(* Logix 5000 project; controller FV vendor 1 type 14 code 217 rev 31.11; software revision 31.00; part 57 of 63 *)
(* tags used below, declared in another part *)
   CWD : CHECKWORD_FLAGS;
   FV_AV1 : PlantItem;   // AV1
   FV_B42 : INT[255];   // YSVCIP_FLG
   FV_B42_0_2_OutputBit : BOOL;
   FV_B52 : INT[255];   // WASTE_FLG
   FV_N141 : INT[255];   // YSV1 DATA
   FV_N142 : INT[255];   // YSV2 DATA
   FV_N143 : INT[255];   // YSV3 DATA
   FV_N40 : INT[255];   // YSVCIP<PC
   FV_N41 : INT[255];   // YSVCIP>PC
   FV_N50 : INT[255];   // WASTE<PC
   FV_N51 : INT[255];   // WASTE>PC
   FV_T43 : TIMER[10];
   FV_T53 : TIMER[10];
   FV_YSV1R : PlantItem;   // YSV1R
   FV_YSV2O : PlantItem;   // YSV2O
   FV_YSV3O : PlantItem;   // YSV3O
(* FV_Common, continued *)

ROUTINE FV_YSVCIP_CP_21   (* ladder *)
   // Reset command interpreter step counter
   0: XIC(S:FS)CLR(FV_N41[16]);
   // RESET
   1: EQU(FV_N41[16],0)MCR();
   2: OTU(FV_B42[0].0);
   3: OTU(FV_B42[0].1);
   4: OTU(FV_B42[0].8);
   5: FLL(0,FV_N41[0],16);
   // Set PCparameter buffer to 'Null' value
   6: FLL(-32768,FV_N40[1],7);
   7: CLR(FV_N40[0]);
   8: MOV(1,FV_N41[16]);
   9: MCR();
   // ALLOW STARTUP DIALOG
   10: EQU(FV_N41[16],1)MCR();
   // Set process status = ready
   11: MOV(1,FV_N41[0]);
   // Allow startup if any vessel is inactive or on storage control only
   12: [[EQU(FV_N141[0],0) ,EQU(FV_N141[0],5) ] ,[EQU(FV_N142[0],0) ,EQU(FV_N142[0],5) ] ,[EQU(FV_N143[0],0) ,EQU(FV_N143[0],5) ] ]OTE(FV_N41[2].0);
   // Advance step if start selected
   13: XIC(FV_N41[2].0)XIC(FV_N40[0].0)MOV(2,FV_N41[16]);
   14: MCR();
   // WAIT FOR STARTUP DIALOG COMPLETE
   15: EQU(FV_N41[16],2)MCR();
   // If YSV1 requested and YSV1 not involved in any other startup dialog set lock flag
   16: EQU(FV_N40[1],1)[EQU(FV_N141[0],0) ,EQU(FV_N141[0],5) ][EQU(FV_N141[4],0) ,XIC(FV_N141[4].3) ]OTE(FV_N141[4].3);
   // If YSV2 requested and YSV2 not involved in any other startup dialog set lock flag
   17: EQU(FV_N40[1],2)[EQU(FV_N142[0],0) ,EQU(FV_N142[0],5) ][EQU(FV_N142[4],0) ,XIC(FV_N142[4].3) ]OTE(FV_N142[4].3);
   // If YSV3 requested and YSV3 not involved in any other startup dialog set lock flag
   18: EQU(FV_N40[1],3)[EQU(FV_N143[0],0) ,EQU(FV_N143[0],5) ][EQU(FV_N143[4],0) ,XIC(FV_N143[4].3) ]OTE(FV_N143[4].3);
   // Allow start confirmed button if selected YSV could be locked
   19: [XIC(FV_N141[4].3) ,XIC(FV_N142[4].3) ,XIC(FV_N143[4].3) ]OTE(FV_N41[2].1);
   // Startup dialog guard timer
   20: TON(FV_T43[0],?,?);
   // Reset command processor if dialog cancel selected or startup dialog timer expired
   21: [XIC(FV_N40[0].15) ,XIC(FV_T43[0].DN) ]CLR(FV_N41[16]);
   // Advance step if start available and selected
   22: XIC(FV_N40[0].1)XIC(FV_N41[2].1)[MOV(3,FV_N41[16]) ,CLR(FV_N40[0]) ];
   23: MCR();
   // COMPLETE STARTUP DIALOG
   24: EQU(FV_N41[16],3)MCR();
   // If YSV 1 selected, set YSV1 status = Cleaning
   25: EQU(FV_N40[1],1)MOV(3,FV_N141[0]);
   // If YSV 2 selected, set YSV2 status =Cleaning
   26: EQU(FV_N40[1],2)MOV(3,FV_N142[0]);
   // If YSV 3 selected, set YSV3 status =Cleaning
   27: EQU(FV_N40[1],3)MOV(3,FV_N143[0]);
   // Set YSV CIP Process Status = Running
   28: MOV(2,FV_N41[0]);
   29: OTL(FV_B42[0].0);
   30: OTL(FV_B42[0].1);
   31: OTL(FV_N41[2].2);
   32: MOV(10,FV_N41[1]);
   33: MOV(10,FV_N41[3]);
   34: MOV(-1,FV_N41[16]);
   35: CLR(FV_N40[0]);
   36: MCR();
   // HANDLE STOP BUTTON
   37: XIC(FV_N40[0].2)XIC(FV_N41[2].2)MCR();
   38: OTU(FV_B42[0].1);
   39: OTU(FV_N41[2].2);
   40: OTL(FV_N41[2].3);
   41: OTL(FV_N41[2].4);
   42: MOV(3,FV_N41[0]);
   43: MOV(0,FV_N41[1]);
   44: CLR(FV_N40[0]);
   45: MCR();
   // HANDLE CONTINUE BUTTON
   46: XIC(FV_N40[0].3)XIC(FV_N41[2].3)MCR();
   47: OTL(FV_B42[0].1);
   48: OTL(FV_N41[2].2);
   49: OTU(FV_N41[2].3);
   // Reset process alarm and parameters
   50: OTU(FV_N41[2].4);
   51: FLL(0,FV_N41[4],4);
   52: MOV(2,FV_N41[0]);
   // Set current Step = Restart Step
   53: MOV(FV_N41[3],FV_N41[1]);
   54: CLR(FV_N40[0]);
   55: MCR();
   // HANDLE ABORT BUTTON
   56: XIC(FV_N40[0].4)XIC(FV_N41[2].4)MCR();
   57: OTU(FV_B42[0].0);
   // Set YSV's operation to no-operation
   58: JSR(FV_Set_FV_Datafile_Value,3,0,FV_N41[15],0);
   59: CLR(FV_N41[16]);
   60: CLR(FV_N40[0]);
   61: MCR();
   // Copy step number for PC to display if running
   62: XIC(FV_B42[0].1)MOV(FV_N41[1],FV_N41[9]);
END_ROUTINE

ROUTINE FV_YSVCIP_MC_20   (* ladder *)
   // Run YSV CIP Command Processor
   0: JSR(FV_YSVCIP_CP_21,0);
   // Run YSV CIP process control program
   1: XIC(FV_B42[0].0)JSR(FV_YSVCIP_PRO_22,0);
   // PostScan YSV CIP control program
   2: XIO(FV_B42[0].0)OSR(FV_B42[0].2,FV_B42_0_2_OutputBit)XIC(FV_B42_0_2_OutputBit)JSR(FV_YSVCIP_PRO_22,0);
END_ROUTINE

ROUTINE FV_YSVCIP_PRO_22   (* ladder *)
   // YSV CIP - STEP 10 - Initialize
   0: XIC(FV_B42[0].1)EQU(FV_N41[1],10)MCR();
   // Set restart step for this process
   1: MOV(10,FV_N41[3]);
   // Make pointer to selected YSV's data file
   2: ADD(FV_N40[1],140,FV_N41[15]);
   // Set rouser to automatic
   3: JSR(FV_Set_FV_Datafile_Value,3,0,FV_N41[15],3);
   // Make pointer to YSV's Attemporation Data File
   4: ADD(FV_N40[1],135,FV_N41[14]);
   // Stop attemporation control on YSV
   5: [JSR(FV_Set_FV_Datafile_Value,3,0,FV_N41[14],24) ,JSR(FV_Set_FV_Datafile_Value,3,0,FV_N41[14],26) JSR(FV_Set_FV_Datafile_Value,3,0,FV_N41[14],27) JSR(FV_Set_FV_Datafile_Value,3,0,FV_N41[14],28) JSR(FV_Set_FV_Datafile_Value,3,0,FV_N41[14],29) ];
   // Advance to next step
   6: MOV(20,FV_N41[1]);
   7: MCR();
   // YSV CIP - STEP 20 - Cleaning Route Open
   8: XIC(FV_B42[0].1)EQU(FV_N41[1],20)MCR();
   // Set restart step for this process
   9: MOV(20,FV_N41[3]);
   // Request inlet / outlet valve on correct vessel
   10: [EQU(FV_N40[1],1) OTE(FV_AV1.DriveBits.3) ,EQU(FV_N40[1],2) OTE(FV_YSV2O.DriveBits.3) ,EQU(FV_N40[1],3) OTE(FV_YSV3O.DriveBits.3) ];
   // Allow operator to select process end button
   11: OTE(FV_N41[2].5);
   // Advance to next step when End selected
   12: XIC(FV_N40[0].5)MOV(30,FV_N41[1]);
   13: MCR();
   // YSV CIP - STEP 30 - Reset YSV
   14: XIC(FV_B42[0].1)EQU(FV_N41[1],30)MCR();
   // Reset Dirty flag on this YSV
   15: JSR(FV_Clear_Flag_In_FV_Datafile,3,FV_N41[15],1,0);
   // Set status of YSV to no-operation
   16: JSR(FV_Set_FV_Datafile_Value,3,0,FV_N41[15],0);
   17: CLR(FV_N41[16]);
   18: MCR();
   // CHECK FOR ALARM CONDITIONS
   19: XIC(FV_B42[0].1)MCR();
   20: EQU(FV_N40[1],1)[XIC(FV_AV1.CW.[CWD.FAULT]) ,XIC(FV_YSV1R.CW.[CWD.FAULT]) ]OTU(FV_B42[0].1);
   21: GRT(FV_N41[4],0)OTU(FV_B42[0].1);
   22: XIO(FV_B42[0].1)[MOV(4,FV_N41[0]) ,OTU(FV_N41[2].2) ,OTL(FV_N41[2].3) ,OTL(FV_N41[2].4) ,MOV(0,FV_N41[1]) ];
   23: MCR();
END_ROUTINE

ROUTINE FV_YSVWSTE_CP_26   (* ladder *)
   // Reset command interpreter step counter
   0: XIC(S:FS)CLR(FV_N51[16]);
   // RESET
   1: EQU(FV_N51[16],0)MCR();
   2: OTU(FV_B52[0].0);
   3: OTU(FV_B52[0].1);
   4: OTU(FV_B52[0].8);
   5: FLL(0,FV_N51[0],16);
   // Set PCparameter buffer to 'Null' value
   6: FLL(-32768,FV_N50[1],7);
   7: CLR(FV_N50[0]);
   8: MOV(1,FV_N51[16]);
   9: MCR();
   // ALLOW STARTUP DIALOG
   10: EQU(FV_N51[16],1)MCR();
   // Set process status = ready
   11: MOV(1,FV_N51[0]);
   // Allow startup if any vessel is inactive or on storage control only
   12: [[EQU(FV_N141[0],0) ,EQU(FV_N141[0],5) ] ,[EQU(FV_N142[0],0) ,EQU(FV_N142[0],5) ] ,[EQU(FV_N143[0],0) ,EQU(FV_N143[0],5) ] ]OTE(FV_N51[2].0);
   // Advance step if start selected
   13: XIC(FV_N51[2].0)XIC(FV_N50[0].0)MOV(2,FV_N51[16]);
   14: MCR();
   // WAIT FOR STARTUP DIALOG COMPLETE
   15: EQU(FV_N51[16],2)MCR();
   // If YSV1 requested and YSV1 not involved in any other startup dialog set lock flag
   16: EQU(FV_N50[1],1)[EQU(FV_N141[0],0) ,EQU(FV_N141[0],5) ][EQU(FV_N141[4],0) ,XIC(FV_N141[4].4) ]OTE(FV_N141[4].4);
   // If YSV2 requested and YSV2 not involved in any other startup dialog set lock flag
   17: EQU(FV_N50[1],2)[EQU(FV_N142[0],0) ,EQU(FV_N142[0],5) ][EQU(FV_N142[4],0) ,XIC(FV_N142[4].4) ]OTE(FV_N142[4].4);
   // If YSV3 requested and YSV3 not involved in any other startup dialog set lock flag
   18: EQU(FV_N50[1],3)[EQU(FV_N143[0],0) ,EQU(FV_N143[0],5) ][EQU(FV_N143[4],0) ,XIC(FV_N143[4].4) ]OTE(FV_N143[4].4);
   // Allow start confirmed button if selected YSV could be locked
   19: [XIC(FV_N141[4].4) ,XIC(FV_N142[4].4) ,XIC(FV_N143[4].4) ]OTE(FV_N51[2].1);
   // Startup dialog guard timer
   20: TON(FV_T53[0],?,?);
   // Reset command processor if dialog cancel selected or startup dialog timer expired
   21: [XIC(FV_N50[0].15) ,XIC(FV_T53[0].DN) ]CLR(FV_N51[16]);
   // Advance step if start available and selected
   22: XIC(FV_N50[0].1)XIC(FV_N51[2].1)[MOV(3,FV_N51[16]) ,CLR(FV_N50[0]) ];
   23: MCR();
   // COMPLETE STARTUP DIALOG
   24: EQU(FV_N51[16],3)MCR();
   // If YSV 1 selected, save YSV1 status
   25: EQU(FV_N50[1],1)MOV(FV_N141[0],FV_N51[13]);
   // If YSV2 selected, save YSV2 status
   26: EQU(FV_N50[1],2)MOV(FV_N142[0],FV_N51[13]);
   // If YSV 3 selected, save YSV3 status
   27: EQU(FV_N50[1],3)MOV(FV_N143[0],FV_N51[13]);
   // If YSV 1 selected, set YSV1 status = Transfer to Waste
   28: EQU(FV_N50[1],1)MOV(4,FV_N141[0]);
   // If YSV 2 selected, set YSV2 status =Transfer to Waste
   29: EQU(FV_N50[1],2)MOV(4,FV_N142[0]);
   // If YSV 3 selected, set YSV3 status = Transfer to Waste
   30: EQU(FV_N50[1],3)MOV(4,FV_N143[0]);
   // Set YSV to Waste Process Status = Running
   31: MOV(2,FV_N51[0]);
